   // stn[25].wipBtn[5,2] := 38000;
   // stn[25].wipBtn[5,3] := 1000;
   // stn[25].wipBtn[5,4] := 1000;
   // stn[25].wipBtn[5,5] := 1000;
   // stn[25].wipBtn[5,6] := 43000;
   // stn[25].wipBtn[5,7] := 37000;
   // stn[25].wipBtn[6,0] := 1000;
   // stn[25].wipBtn[6,1] := 244000;
   // stn[25].wipBtn[6,2] := 46000;
   // stn[25].wipBtn[6,3] := 1000;
   // stn[25].wipBtn[6,4] := 1000;
   // stn[25].wipBtn[6,5] := 1000;
   // stn[25].wipBtn[6,6] := 43000;
   // stn[25].wipBtn[6,7] := 37000;
   // stn[25].wipBtn[7,0] := 1000;
   // stn[25].wipBtn[7,1] := 244000;
   // stn[25].wipBtn[7,2] := 44000;
   // stn[25].wipBtn[7,3] := 1000;
   // stn[25].wipBtn[7,4] := 1000;
   // stn[25].wipBtn[7,5] := 1000;
   // stn[25].wipBtn[7,6] := 39000;
   // stn[25].wipBtn[7,7] := 45000;
   // stn[25].wipBtn[8,0] := 1000;
   // stn[25].wipBtn[8,1] := 244000;
   // stn[25].wipBtn[8,2] := 52000;
   // stn[25].wipBtn[8,3] := 1000;
   // stn[25].wipBtn[8,4] := 1000;
   // stn[25].wipBtn[8,5] := 1000;
   // stn[25].wipBtn[8,6] := 26000;
   // stn[25].wipBtn[8,7] := 19000;
   // stn[25].wipBtn[9,0] := 1000;
   // stn[25].wipBtn[9,1] := 244000;
   // stn[25].wipBtn[9,2] := 53000;
   // stn[25].wipBtn[9,3] := 1000;
   // stn[25].wipBtn[9,4] := 1000;
   // stn[25].wipBtn[9,5] := 1000;
   // stn[25].wipBtn[9,6] := 32000;
   // stn[25].wipBtn[9,7] := 74000;
   // stn[25].wipBtn[10,0] := 1000;
   // stn[25].wipBtn[10,1] := 244000;
   // stn[25].wipBtn[10,2] := 54000;
   // stn[25].wipBtn[10,3] := 1000;
   // stn[25].wipBtn[10,4] := 1000;
   // stn[25].wipBtn[10,5] := 1000;
   // stn[25].wipBtn[10,6] := 32000;
   // stn[25].wipBtn[10,7] := 72000;
   // stn[25].wipBtn[11,0] := 1000;
   // stn[25].wipBtn[11,1] := 244000;
   // stn[25].wipBtn[11,2] := 58000;
   // stn[25].wipBtn[11,3] := 1000;
   // stn[25].wipBtn[11,4] := 1000;
   // stn[25].wipBtn[11,5] := 1000;
   // stn[25].wipBtn[11,6] := 26000;
   // stn[25].wipBtn[11,7] := 19000;
   // stn[25].wipBtn[12,0] := 1000;
   // stn[25].wipBtn[12,1] := 244000;
   // stn[25].wipBtn[12,2] := 85000;
   // stn[25].wipBtn[12,3] := 1000;
   // stn[25].wipBtn[12,4] := 1000;
   // stn[25].wipBtn[12,5] := 1000;
   // stn[25].wipBtn[12,6] := 32000;
   // stn[25].wipBtn[12,7] := 72000;
   // stn[25].wipBtn[13,0] := 1000;
   // stn[25].wipBtn[13,1] := 244000;
   // stn[25].wipBtn[13,2] := 99000;
   // stn[25].wipBtn[13,3] := 1000;
   // stn[25].wipBtn[13,4] := 1000;
   // stn[25].wipBtn[13,5] := 1000;
   // stn[25].wipBtn[13,6] := 39000;
   // stn[25].wipBtn[13,7] := 45000;
   // stn[25].wipBtn[14,0] := 1000;
   // stn[25].wipBtn[14,1] := 244000;
   // stn[25].wipBtn[14,2] := 100000;
   // stn[25].wipBtn[14,3] := 1000;
   // stn[25].wipBtn[14,4] := 1000;
   // stn[25].wipBtn[14,5] := 1000;
   // stn[25].wipBtn[14,6] := 43000;
   // stn[25].wipBtn[14,7] := 37000;
   // stn[25].wipBtn[15,0] := 1000;
   // stn[25].wipBtn[15,1] := 244000;
   // stn[25].wipBtn[15,2] := 100000;
   // stn[25].wipBtn[15,3] := 1000;
   // stn[25].wipBtn[15,4] := 1000;
   // stn[25].wipBtn[15,5] := 1000;
   // stn[25].wipBtn[15,6] := 36000;
   // stn[25].wipBtn[15,7] := 37000;
   // stn[25].wipBtn[16,0] := 1000;
   // stn[25].wipBtn[16,1] := 244000;
   // stn[25].wipBtn[16,2] := 218000;
   // stn[25].wipBtn[16,3] := 1000;
   // stn[25].wipBtn[16,4] := 1000;
   // stn[25].wipBtn[16,5] := 1000;
   // stn[25].wipBtn[16,6] := 219000;
   // stn[25].wipBtn[16,7] := 224000;
   // stn[25].wipBtn[17,0] := 1000;
   // stn[25].wipBtn[17,1] := 244000;
   // stn[25].wipBtn[17,2] := 198000;
   // stn[25].wipBtn[17,3] := 1000;
   // stn[25].wipBtn[17,4] := 1000;
   // stn[25].wipBtn[17,5] := 1000;
   // stn[25].wipBtn[17,6] := 220000;
   // stn[25].wipBtn[17,7] := 223000;
   // stn[25].wipBtn[18,0] := 1000;
   // stn[25].wipBtn[18,1] := 244000;
   // stn[25].wipBtn[18,2] := 199000;
   // stn[25].wipBtn[18,3] := 1000;
   // stn[25].wipBtn[18,4] := 1000;
   // stn[25].wipBtn[18,5] := 1000;
   // stn[25].wipBtn[18,6] := 219000;
   // stn[25].wipBtn[18,7] := 224000;
   // stn[25].wipBtn[19,0] := 1000;
   // stn[25].wipBtn[19,1] := 244000;
   // stn[25].wipBtn[19,2] := 225000;
   // stn[25].wipBtn[19,3] := 1000;
   // stn[25].wipBtn[19,4] := 1000;
   // stn[25].wipBtn[19,5] := 1000;
   // stn[25].wipBtn[19,6] := 226000;
   // stn[25].wipBtn[19,7] := 227000;
   // stn[25].wipBtn[20,0] := 1000;
   // stn[25].wipBtn[20,1] := 244000;
   // stn[25].wipBtn[20,2] := 18000;
   // stn[25].wipBtn[20,3] := 1000;
   // stn[25].wipBtn[20,4] := 1000;
   // stn[25].wipBtn[20,5] := 1000;
   // stn[25].wipBtn[20,6] := 25000;
   // stn[25].wipBtn[20,7] := 17000;
   // stn[25].wipBtn[21,0] := 1000;
   // stn[25].wipBtn[21,1] := 244000;
   // stn[25].wipBtn[21,2] := 1000;
   // stn[25].wipBtn[21,3] := 32000;
   // stn[25].wipBtn[21,4] := 1000;
   // stn[25].wipBtn[21,5] := 1000;
   // stn[25].wipBtn[21,6] := 51000;
   // stn[25].wipBtn[21,7] := 31000;
   // stn[25].wipBtn[22,0] := 1000;
   // stn[25].wipBtn[22,1] := 244000;
   // stn[25].wipBtn[22,2] := 1000;
   // stn[25].wipBtn[22,3] := 220000;
   // stn[25].wipBtn[22,4] := 1000;
   // stn[25].wipBtn[22,5] := 1000;
   // stn[25].wipBtn[22,6] := 222000;
   // stn[25].wipBtn[22,7] := 223000;
   // stn[25].wipBtn[23,0] := 1000;
   // stn[25].wipBtn[23,1] := 244000;
   // stn[25].wipBtn[23,2] := 221000;
   // stn[25].wipBtn[23,3] := 1000;
   // stn[25].wipBtn[23,4] := 1000;
   // stn[25].wipBtn[23,5] := 1000;
   // stn[25].wipBtn[23,6] := 220000;
   // stn[25].wipBtn[23,7] := 223000;
   // stn[25].wipBtn[24,0] := 1000;
   // stn[25].wipBtn[24,1] := 1000;
   // stn[25].wipBtn[24,2] := 1000;
   // stn[25].wipBtn[24,3] := 1000;
   // stn[25].wipBtn[24,4] := 1000;
   // stn[25].wipBtn[24,5] := 1000;
   // stn[25].wipBtn[24,6] := 1000;
   // stn[25].wipBtn[24,7] := 1000;
   // stn[25].wipBtn[25,0] := 1000;
   // stn[25].wipBtn[25,1] := 1000;
   // stn[25].wipBtn[25,2] := 1000;
   // stn[25].wipBtn[25,3] := 1000;
   // stn[25].wipBtn[25,4] := 1000;
   // stn[25].wipBtn[25,5] := 1000;
   // stn[25].wipBtn[25,6] := 1000;
   // stn[25].wipBtn[25,7] := 1000;
   // stn[25].wipBtn[26,0] := 1000;
   // stn[25].wipBtn[26,1] := 1000;
   // stn[25].wipBtn[26,2] := 1000;
   // stn[25].wipBtn[26,3] := 1000;
   // stn[25].wipBtn[26,4] := 1000;
   // stn[25].wipBtn[26,5] := 1000;
   // stn[25].wipBtn[26,6] := 1000;
   // stn[25].wipBtn[26,7] := 1000;
   // stn[25].wipBtn[27,0] := 1000;
   // stn[25].wipBtn[27,1] := 1000;
   // stn[25].wipBtn[27,2] := 1000;
   // stn[25].wipBtn[27,3] := 1000;
   // stn[25].wipBtn[27,4] := 1000;
   // stn[25].wipBtn[27,5] := 1000;
   // stn[25].wipBtn[27,6] := 1000;
   // stn[25].wipBtn[27,7] := 1000;
   // stn[25].wipBtn[28,0] := 1000;
   // stn[25].wipBtn[28,1] := 1000;
   // stn[25].wipBtn[28,2] := 1000;
   // stn[25].wipBtn[28,3] := 1000;
   // stn[25].wipBtn[28,4] := 1000;
   // stn[25].wipBtn[28,5] := 1000;
   // stn[25].wipBtn[28,6] := 1000;
   // stn[25].wipBtn[28,7] := 1000;
   // stn[25].wipBtn[29,0] := 1000;
   // stn[25].wipBtn[29,1] := 1000;
   // stn[25].wipBtn[29,2] := 1000;
   // stn[25].wipBtn[29,3] := 1000;
   // stn[25].wipBtn[29,4] := 1000;
   // stn[25].wipBtn[29,5] := 1000;
   // stn[25].wipBtn[29,6] := 1000;
   // stn[25].wipBtn[29,7] := 1000;
   // stn[25].wipBtn[30,0] := 1000;
   // stn[25].wipBtn[30,1] := 1000;
   // stn[25].wipBtn[30,2] := 1000;
   // stn[25].wipBtn[30,3] := 1000;
   // stn[25].wipBtn[30,4] := 1000;
   // stn[25].wipBtn[30,5] := 1000;
   // stn[25].wipBtn[30,6] := 1000;
   // stn[25].wipBtn[30,7] := 1000;
   // stn[25].wipBtn[31,0] := 1000;
   // stn[25].wipBtn[31,1] := 1000;
   // stn[25].wipBtn[31,2] := 1000;
   // stn[25].wipBtn[31,3] := 1000;
   // stn[25].wipBtn[31,4] := 1000;
   // stn[25].wipBtn[31,5] := 1000;
   // stn[25].wipBtn[31,6] := 1000;
   // stn[25].wipBtn[31,7] := 1000;
   // stn[25].wipBtn[32,0] := 1000;
   // stn[25].wipBtn[32,1] := 1000;
   // stn[25].wipBtn[32,2] := 1000;
   // stn[25].wipBtn[32,3] := 1000;
   // stn[25].wipBtn[32,4] := 1000;
   // stn[25].wipBtn[32,5] := 1000;
   // stn[25].wipBtn[32,6] := 1000;
   // stn[25].wipBtn[32,7] := 1000;
   // stn[25].wipBtn[33,0] := 1000;
   // stn[25].wipBtn[33,1] := 1000;
   // stn[25].wipBtn[33,2] := 1000;
   // stn[25].wipBtn[33,3] := 1000;
   // stn[25].wipBtn[33,4] := 1000;
   // stn[25].wipBtn[33,5] := 1000;
   // stn[25].wipBtn[33,6] := 1000;
   // stn[25].wipBtn[33,7] := 1000;
   // stn[25].wipBtn[34,0] := 1000;
   // stn[25].wipBtn[34,1] := 1000;
   // stn[25].wipBtn[34,2] := 1000;
   // stn[25].wipBtn[34,3] := 1000;
   // stn[25].wipBtn[34,4] := 1000;
   // stn[25].wipBtn[34,5] := 1000;
   // stn[25].wipBtn[34,6] := 1000;
   // stn[25].wipBtn[34,7] := 1000;
   // stn[25].wipBtn[35,0] := 1000;
   // stn[25].wipBtn[35,1] := 1000;
   // stn[25].wipBtn[35,2] := 1000;
   // stn[25].wipBtn[35,3] := 1000;
   // stn[25].wipBtn[35,4] := 1000;
   // stn[25].wipBtn[35,5] := 1000;
   // stn[25].wipBtn[35,6] := 1000;
   // stn[25].wipBtn[35,7] := 1000;
   // stn[25].wipBtn[36,0] := 1000;
   // stn[25].wipBtn[36,1] := 1000;
   // stn[25].wipBtn[36,2] := 1000;
   // stn[25].wipBtn[36,3] := 1000;
   // stn[25].wipBtn[36,4] := 1000;
   // stn[25].wipBtn[36,5] := 1000;
   // stn[25].wipBtn[36,6] := 1000;
   // stn[25].wipBtn[36,7] := 1000;
   // stn[25].wipBtn[37,0] := 1000;
   // stn[25].wipBtn[37,1] := 1000;
   // stn[25].wipBtn[37,2] := 1000;
   // stn[25].wipBtn[37,3] := 1000;
   // stn[25].wipBtn[37,4] := 1000;
   // stn[25].wipBtn[37,5] := 1000;
   // stn[25].wipBtn[37,6] := 1000;
   // stn[25].wipBtn[37,7] := 1000;
   // stn[25].wipBtn[38,0] := 1000;
   // stn[25].wipBtn[38,1] := 1000;
   // stn[25].wipBtn[38,2] := 1000;
   // stn[25].wipBtn[38,3] := 1000;
   // stn[25].wipBtn[38,4] := 1000;
   // stn[25].wipBtn[38,5] := 1000;
   // stn[25].wipBtn[38,6] := 1000;
   // stn[25].wipBtn[38,7] := 1000;
   // stn[25].wipBtn[39,0] := 1000;
   // stn[25].wipBtn[39,1] := 1000;
   // stn[25].wipBtn[39,2] := 1000;
   // stn[25].wipBtn[39,3] := 1000;
   // stn[25].wipBtn[39,4] := 1000;
   // stn[25].wipBtn[39,5] := 1000;
   // stn[25].wipBtn[39,6] := 1000;
   // stn[25].wipBtn[39,7] := 1000;
   // stn[25].wipBtn[40,0] := 1000;
   // stn[25].wipBtn[40,1] := 1000;
   // stn[25].wipBtn[40,2] := 1000;
   // stn[25].wipBtn[40,3] := 1000;
   // stn[25].wipBtn[40,4] := 1000;
   // stn[25].wipBtn[40,5] := 1000;
   // stn[25].wipBtn[40,6] := 1000;
   // stn[25].wipBtn[40,7] := 1000;
   // stn[25].wipBtn[41,0] := 1000;
   // stn[25].wipBtn[41,1] := 1000;
   // stn[25].wipBtn[41,2] := 1000;
   // stn[25].wipBtn[41,3] := 1000;
   // stn[25].wipBtn[41,4] := 1000;
   // stn[25].wipBtn[41,5] := 1000;
   // stn[25].wipBtn[41,6] := 1000;
   // stn[25].wipBtn[41,7] := 1000;
   // stn[25].wipBtn[42,0] := 1000;
   // stn[25].wipBtn[42,1] := 1000;
   // stn[25].wipBtn[42,2] := 1000;
   // stn[25].wipBtn[42,3] := 1000;
   // stn[25].wipBtn[42,4] := 1000;
   // stn[25].wipBtn[42,5] := 1000;
   // stn[25].wipBtn[42,6] := 1000;
   // stn[25].wipBtn[42,7] := 1000;
   // stn[25].wipBtn[43,0] := 1000;
   // stn[25].wipBtn[43,1] := 1000;
   // stn[25].wipBtn[43,2] := 1000;
   // stn[25].wipBtn[43,3] := 1000;
   // stn[25].wipBtn[43,4] := 1000;
   // stn[25].wipBtn[43,5] := 1000;
   // stn[25].wipBtn[43,6] := 1000;
   // stn[25].wipBtn[43,7] := 1000;
   // stn[25].wipBtn[44,0] := 1000;
   // stn[25].wipBtn[44,1] := 1000;
   // stn[25].wipBtn[44,2] := 1000;
   // stn[25].wipBtn[44,3] := 1000;
   // stn[25].wipBtn[44,4] := 1000;
   // stn[25].wipBtn[44,5] := 1000;
   // stn[25].wipBtn[44,6] := 1000;
   // stn[25].wipBtn[44,7] := 1000;
   // stn[25].wipBtn[45,0] := 1000;
   // stn[25].wipBtn[45,1] := 1000;
   // stn[25].wipBtn[45,2] := 1000;
   // stn[25].wipBtn[45,3] := 1000;
   // stn[25].wipBtn[45,4] := 1000;
   // stn[25].wipBtn[45,5] := 1000;
   // stn[25].wipBtn[45,6] := 1000;
   // stn[25].wipBtn[45,7] := 1000;
   // stn[25].wipBtn[46,0] := 1000;
   // stn[25].wipBtn[46,1] := 1000;
   // stn[25].wipBtn[46,2] := 1000;
   // stn[25].wipBtn[46,3] := 1000;
   // stn[25].wipBtn[46,4] := 1000;
   // stn[25].wipBtn[46,5] := 1000;
   // stn[25].wipBtn[46,6] := 1000;
   // stn[25].wipBtn[46,7] := 1000;
   // stn[25].wipBtn[47,0] := 1000;
   // stn[25].wipBtn[47,1] := 1000;
   // stn[25].wipBtn[47,2] := 1000;
   // stn[25].wipBtn[47,3] := 1000;
   // stn[25].wipBtn[47,4] := 1000;
   // stn[25].wipBtn[47,5] := 1000;
   // stn[25].wipBtn[47,6] := 1000;
   // stn[25].wipBtn[47,7] := 1000;
   // stn[25].wipBtn[48,0] := 1000;
   // stn[25].wipBtn[48,1] := 1000;
   // stn[25].wipBtn[48,2] := 1000;
   // stn[25].wipBtn[48,3] := 1000;
   // stn[25].wipBtn[48,4] := 1000;
   // stn[25].wipBtn[48,5] := 1000;
   // stn[25].wipBtn[48,6] := 1000;
   // stn[25].wipBtn[48,7] := 1000;
   // stn[25].wipBtn[49,0] := 1000;
   // stn[25].wipBtn[49,1] := 1000;
   // stn[25].wipBtn[49,2] := 1000;
   // stn[25].wipBtn[49,3] := 1000;
   // stn[25].wipBtn[49,4] := 1000;
   // stn[25].wipBtn[49,5] := 1000;
   // stn[25].wipBtn[49,6] := 1000;
   // stn[25].wipBtn[49,7] := 1000;
   // stn[26].wipBtn[0,0] := 1000;
   // stn[26].wipBtn[0,1] := 244000;
   // stn[26].wipBtn[0,2] := 46000;
   // stn[26].wipBtn[0,3] := 1000;
   // stn[26].wipBtn[0,4] := 1000;
   // stn[26].wipBtn[0,5] := 1000;
   // stn[26].wipBtn[0,6] := 43000;
   // stn[26].wipBtn[0,7] := 37000;
   // stn[26].wipBtn[1,0] := 1000;
   // stn[26].wipBtn[1,1] := 244000;
   // stn[26].wipBtn[1,2] := 100000;
   // stn[26].wipBtn[1,3] := 1000;
   // stn[26].wipBtn[1,4] := 1000;
   // stn[26].wipBtn[1,5] := 1000;
   // stn[26].wipBtn[1,6] := 43000;
   // stn[26].wipBtn[1,7] := 37000;
   // stn[26].wipBtn[2,0] := 1000;
   // stn[26].wipBtn[2,1] := 244000;
   // stn[26].wipBtn[2,2] := 100000;
   // stn[26].wipBtn[2,3] := 1000;
   // stn[26].wipBtn[2,4] := 1000;
   // stn[26].wipBtn[2,5] := 1000;
   // stn[26].wipBtn[2,6] := 36000;
   // stn[26].wipBtn[2,7] := 37000;
   // stn[26].wipBtn[3,0] := 1000;
   // stn[26].wipBtn[3,1] := 244000;
   // stn[26].wipBtn[3,2] := 15000;
   // stn[26].wipBtn[3,3] := 1000;
   // stn[26].wipBtn[3,4] := 1000;
   // stn[26].wipBtn[3,5] := 16000;
   // stn[26].wipBtn[3,6] := 24000;
   // stn[26].wipBtn[3,7] := 14000;
   // stn[26].wipBtn[4,0] := 1000;
   // stn[26].wipBtn[4,1] := 244000;
   // stn[26].wipBtn[4,2] := 15000;
   // stn[26].wipBtn[4,3] := 14000;
   // stn[26].wipBtn[4,4] := 1000;
   // stn[26].wipBtn[4,5] := 48000;
   // stn[26].wipBtn[4,6] := 34000;
   // stn[26].wipBtn[4,7] := 33000;
   // stn[26].wipBtn[5,0] := 1000;
   // stn[26].wipBtn[5,1] := 244000;
   // stn[26].wipBtn[5,2] := 15000;
   // stn[26].wipBtn[5,3] := 1000;
   // stn[26].wipBtn[5,4] := 1000;
   // stn[26].wipBtn[5,5] := 16000;
   // stn[26].wipBtn[5,6] := 34000;
   // stn[26].wipBtn[5,7] := 14000;
   // stn[26].wipBtn[6,0] := 1000;
   // stn[26].wipBtn[6,1] := 244000;
   // stn[26].wipBtn[6,2] := 71000;
   // stn[26].wipBtn[6,3] := 74000;
   // stn[26].wipBtn[6,4] := 1000;
   // stn[26].wipBtn[6,5] := 59000;
   // stn[26].wipBtn[6,6] := 42000;
   // stn[26].wipBtn[6,7] := 73000;
   // stn[26].wipBtn[7,0] := 1000;
   // stn[26].wipBtn[7,1] := 244000;
   // stn[26].wipBtn[7,2] := 229000;
   // stn[26].wipBtn[7,3] := 232000;
   // stn[26].wipBtn[7,4] := 1000;
   // stn[26].wipBtn[7,5] := 230000;
   // stn[26].wipBtn[7,6] := 228000;
   // stn[26].wipBtn[7,7] := 231000;
   // stn[26].wipBtn[8,0] := 1000;
   // stn[26].wipBtn[8,1] := 244000;
   // stn[26].wipBtn[8,2] := 234000;
   // stn[26].wipBtn[8,3] := 1000;
   // stn[26].wipBtn[8,4] := 1000;
   // stn[26].wipBtn[8,5] := 230000;
   // stn[26].wipBtn[8,6] := 233000;
   // stn[26].wipBtn[8,7] := 232000;
   // stn[26].wipBtn[9,0] := 1000;
   // stn[26].wipBtn[9,1] := 244000;
   // stn[26].wipBtn[9,2] := 237000;
   // stn[26].wipBtn[9,3] := 1000;
   // stn[26].wipBtn[9,4] := 1000;
   // stn[26].wipBtn[9,5] := 238000;
   // stn[26].wipBtn[9,6] := 235000;
   // stn[26].wipBtn[9,7] := 236000;
   // stn[26].wipBtn[10,0] := 1000;
   // stn[26].wipBtn[10,1] := 244000;
   // stn[26].wipBtn[10,2] := 165000;
   // stn[26].wipBtn[10,3] := 1000;
   // stn[26].wipBtn[10,4] := 1000;
   // stn[26].wipBtn[10,5] := 166000;
   // stn[26].wipBtn[10,6] := 235000;
   // stn[26].wipBtn[10,7] := 236000;
   // stn[26].wipBtn[11,0] := 1000;
   // stn[26].wipBtn[11,1] := 244000;
   // stn[26].wipBtn[11,2] := 202000;
   // stn[26].wipBtn[11,3] := 1000;
   // stn[26].wipBtn[11,4] := 1000;
   // stn[26].wipBtn[11,5] := 201000;
   // stn[26].wipBtn[11,6] := 235000;
   // stn[26].wipBtn[11,7] := 236000;
   // stn[26].wipBtn[12,0] := 1000;
   // stn[26].wipBtn[12,1] := 244000;
   // stn[26].wipBtn[12,2] := 241000;
   // stn[26].wipBtn[12,3] := 1000;
   // stn[26].wipBtn[12,4] := 1000;
   // stn[26].wipBtn[12,5] := 242000;
   // stn[26].wipBtn[12,6] := 239000;
   // stn[26].wipBtn[12,7] := 240000;
   // stn[26].wipBtn[13,0] := 1000;
   // stn[26].wipBtn[13,1] := 244000;
   // stn[26].wipBtn[13,2] := 71000;
   // stn[26].wipBtn[13,3] := 73000;
   // stn[26].wipBtn[13,4] := 1000;
   // stn[26].wipBtn[13,5] := 59000;
   // stn[26].wipBtn[13,6] := 34000;
   // stn[26].wipBtn[13,7] := 74000;
   // stn[26].wipBtn[14,0] := 1000;
   // stn[26].wipBtn[14,1] := 1000;
   // stn[26].wipBtn[14,2] := 1000;
   // stn[26].wipBtn[14,3] := 1000;
   // stn[26].wipBtn[14,4] := 1000;
   // stn[26].wipBtn[14,5] := 1000;
   // stn[26].wipBtn[14,6] := 1000;
   // stn[26].wipBtn[14,7] := 1000;
   // stn[26].wipBtn[15,0] := 1000;
   // stn[26].wipBtn[15,1] := 1000;
   // stn[26].wipBtn[15,2] := 1000;
   // stn[26].wipBtn[15,3] := 1000;
   // stn[26].wipBtn[15,4] := 1000;
   // stn[26].wipBtn[15,5] := 1000;
   // stn[26].wipBtn[15,6] := 1000;
   // stn[26].wipBtn[15,7] := 1000;
   // stn[26].wipBtn[16,0] := 1000;
   // stn[26].wipBtn[16,1] := 1000;
   // stn[26].wipBtn[16,2] := 1000;
   // stn[26].wipBtn[16,3] := 1000;
   // stn[26].wipBtn[16,4] := 1000;
   // stn[26].wipBtn[16,5] := 1000;
   // stn[26].wipBtn[16,6] := 1000;
   // stn[26].wipBtn[16,7] := 1000;
   // stn[26].wipBtn[17,0] := 1000;
   // stn[26].wipBtn[17,1] := 1000;
   // stn[26].wipBtn[17,2] := 1000;
   // stn[26].wipBtn[17,3] := 1000;
   // stn[26].wipBtn[17,4] := 1000;
   // stn[26].wipBtn[17,5] := 1000;
   // stn[26].wipBtn[17,6] := 1000;
   // stn[26].wipBtn[17,7] := 1000;
   // stn[26].wipBtn[18,0] := 1000;
   // stn[26].wipBtn[18,1] := 1000;
   // stn[26].wipBtn[18,2] := 1000;
   // stn[26].wipBtn[18,3] := 1000;
   // stn[26].wipBtn[18,4] := 1000;
   // stn[26].wipBtn[18,5] := 1000;
   // stn[26].wipBtn[18,6] := 1000;
   // stn[26].wipBtn[18,7] := 1000;
   // stn[26].wipBtn[19,0] := 1000;
   // stn[26].wipBtn[19,1] := 1000;
   // stn[26].wipBtn[19,2] := 1000;
   // stn[26].wipBtn[19,3] := 1000;
   // stn[26].wipBtn[19,4] := 1000;
   // stn[26].wipBtn[19,5] := 1000;
   // stn[26].wipBtn[19,6] := 1000;
   // stn[26].wipBtn[19,7] := 1000;
   // stn[26].wipBtn[20,0] := 1000;
   // stn[26].wipBtn[20,1] := 1000;
   // stn[26].wipBtn[20,2] := 1000;
   // stn[26].wipBtn[20,3] := 1000;
   // stn[26].wipBtn[20,4] := 1000;
   // stn[26].wipBtn[20,5] := 1000;
   // stn[26].wipBtn[20,6] := 1000;
   // stn[26].wipBtn[20,7] := 1000;
   // stn[26].wipBtn[21,0] := 1000;
   // stn[26].wipBtn[21,1] := 1000;
   // stn[26].wipBtn[21,2] := 1000;
   // stn[26].wipBtn[21,3] := 1000;
   // stn[26].wipBtn[21,4] := 1000;
   // stn[26].wipBtn[21,5] := 1000;
   // stn[26].wipBtn[21,6] := 1000;
   // stn[26].wipBtn[21,7] := 1000;
   // stn[26].wipBtn[22,0] := 1000;
   // stn[26].wipBtn[22,1] := 1000;
   // stn[26].wipBtn[22,2] := 1000;
   // stn[26].wipBtn[22,3] := 1000;
   // stn[26].wipBtn[22,4] := 1000;
   // stn[26].wipBtn[22,5] := 1000;
   // stn[26].wipBtn[22,6] := 1000;
   // stn[26].wipBtn[22,7] := 1000;
   // stn[26].wipBtn[23,0] := 1000;
   // stn[26].wipBtn[23,1] := 1000;
   // stn[26].wipBtn[23,2] := 1000;
   // stn[26].wipBtn[23,3] := 1000;
   // stn[26].wipBtn[23,4] := 1000;
   // stn[26].wipBtn[23,5] := 1000;
   // stn[26].wipBtn[23,6] := 1000;
   // stn[26].wipBtn[23,7] := 1000;
   // stn[26].wipBtn[24,0] := 1000;
   // stn[26].wipBtn[24,1] := 1000;
   // stn[26].wipBtn[24,2] := 1000;
   // stn[26].wipBtn[24,3] := 1000;
   // stn[26].wipBtn[24,4] := 1000;
   // stn[26].wipBtn[24,5] := 1000;
   // stn[26].wipBtn[24,6] := 1000;
   // stn[26].wipBtn[24,7] := 1000;
   // stn[26].wipBtn[25,0] := 1000;
   // stn[26].wipBtn[25,1] := 1000;
   // stn[26].wipBtn[25,2] := 1000;
   // stn[26].wipBtn[25,3] := 1000;
   // stn[26].wipBtn[25,4] := 1000;
   // stn[26].wipBtn[25,5] := 1000;
   // stn[26].wipBtn[25,6] := 1000;
   // stn[26].wipBtn[25,7] := 1000;
   // stn[26].wipBtn[26,0] := 1000;
   // stn[26].wipBtn[26,1] := 1000;
   // stn[26].wipBtn[26,2] := 1000;
   // stn[26].wipBtn[26,3] := 1000;
   // stn[26].wipBtn[26,4] := 1000;
   // stn[26].wipBtn[26,5] := 1000;
   // stn[26].wipBtn[26,6] := 1000;
   // stn[26].wipBtn[26,7] := 1000;
   // stn[26].wipBtn[27,0] := 1000;
   // stn[26].wipBtn[27,1] := 1000;
   // stn[26].wipBtn[27,2] := 1000;
   // stn[26].wipBtn[27,3] := 1000;
   // stn[26].wipBtn[27,4] := 1000;
   // stn[26].wipBtn[27,5] := 1000;
   // stn[26].wipBtn[27,6] := 1000;
   // stn[26].wipBtn[27,7] := 1000;
   // stn[26].wipBtn[28,0] := 1000;
   // stn[26].wipBtn[28,1] := 1000;
   // stn[26].wipBtn[28,2] := 1000;
   // stn[26].wipBtn[28,3] := 1000;
   // stn[26].wipBtn[28,4] := 1000;
   // stn[26].wipBtn[28,5] := 1000;
   // stn[26].wipBtn[28,6] := 1000;
   // stn[26].wipBtn[28,7] := 1000;
   // stn[26].wipBtn[29,0] := 1000;
   // stn[26].wipBtn[29,1] := 1000;
   // stn[26].wipBtn[29,2] := 1000;
   // stn[26].wipBtn[29,3] := 1000;
   // stn[26].wipBtn[29,4] := 1000;
   // stn[26].wipBtn[29,5] := 1000;
   // stn[26].wipBtn[29,6] := 1000;
   // stn[26].wipBtn[29,7] := 1000;
   // stn[26].wipBtn[30,0] := 1000;
   // stn[26].wipBtn[30,1] := 1000;
   // stn[26].wipBtn[30,2] := 1000;
   // stn[26].wipBtn[30,3] := 1000;
   // stn[26].wipBtn[30,4] := 1000;
   // stn[26].wipBtn[30,5] := 1000;
   // stn[26].wipBtn[30,6] := 1000;
   // stn[26].wipBtn[30,7] := 1000;
   // stn[26].wipBtn[31,0] := 1000;
   // stn[26].wipBtn[31,1] := 1000;
   // stn[26].wipBtn[31,2] := 1000;
   // stn[26].wipBtn[31,3] := 1000;
   // stn[26].wipBtn[31,4] := 1000;
   // stn[26].wipBtn[31,5] := 1000;
   // stn[26].wipBtn[31,6] := 1000;
   // stn[26].wipBtn[31,7] := 1000;
   // stn[26].wipBtn[32,0] := 1000;
   // stn[26].wipBtn[32,1] := 1000;
   // stn[26].wipBtn[32,2] := 1000;
   // stn[26].wipBtn[32,3] := 1000;
   // stn[26].wipBtn[32,4] := 1000;
   // stn[26].wipBtn[32,5] := 1000;
   // stn[26].wipBtn[32,6] := 1000;
   // stn[26].wipBtn[32,7] := 1000;
   // stn[26].wipBtn[33,0] := 1000;
   // stn[26].wipBtn[33,1] := 1000;
   // stn[26].wipBtn[33,2] := 1000;
   // stn[26].wipBtn[33,3] := 1000;
   // stn[26].wipBtn[33,4] := 1000;
   // stn[26].wipBtn[33,5] := 1000;
   // stn[26].wipBtn[33,6] := 1000;
   // stn[26].wipBtn[33,7] := 1000;
   // stn[26].wipBtn[34,0] := 1000;
   // stn[26].wipBtn[34,1] := 1000;
   // stn[26].wipBtn[34,2] := 1000;
   // stn[26].wipBtn[34,3] := 1000;
   // stn[26].wipBtn[34,4] := 1000;
   // stn[26].wipBtn[34,5] := 1000;
   // stn[26].wipBtn[34,6] := 1000;
   // stn[26].wipBtn[34,7] := 1000;
   // stn[26].wipBtn[35,0] := 1000;
   // stn[26].wipBtn[35,1] := 1000;
   // stn[26].wipBtn[35,2] := 1000;
   // stn[26].wipBtn[35,3] := 1000;
   // stn[26].wipBtn[35,4] := 1000;
   // stn[26].wipBtn[35,5] := 1000;
   // stn[26].wipBtn[35,6] := 1000;
   // stn[26].wipBtn[35,7] := 1000;
   // stn[26].wipBtn[36,0] := 1000;
   // stn[26].wipBtn[36,1] := 1000;
   // stn[26].wipBtn[36,2] := 1000;
   // stn[26].wipBtn[36,3] := 1000;
   // stn[26].wipBtn[36,4] := 1000;
   // stn[26].wipBtn[36,5] := 1000;
   // stn[26].wipBtn[36,6] := 1000;
   // stn[26].wipBtn[36,7] := 1000;
   // stn[26].wipBtn[37,0] := 1000;
   // stn[26].wipBtn[37,1] := 1000;
   // stn[26].wipBtn[37,2] := 1000;
   // stn[26].wipBtn[37,3] := 1000;
   // stn[26].wipBtn[37,4] := 1000;
   // stn[26].wipBtn[37,5] := 1000;
   // stn[26].wipBtn[37,6] := 1000;
   // stn[26].wipBtn[37,7] := 1000;
   // stn[26].wipBtn[38,0] := 1000;
   // stn[26].wipBtn[38,1] := 1000;
   // stn[26].wipBtn[38,2] := 1000;
   // stn[26].wipBtn[38,3] := 1000;
   // stn[26].wipBtn[38,4] := 1000;
   // stn[26].wipBtn[38,5] := 1000;
   // stn[26].wipBtn[38,6] := 1000;
   // stn[26].wipBtn[38,7] := 1000;
   // stn[26].wipBtn[39,0] := 1000;
   // stn[26].wipBtn[39,1] := 1000;
   // stn[26].wipBtn[39,2] := 1000;
   // stn[26].wipBtn[39,3] := 1000;
   // stn[26].wipBtn[39,4] := 1000;
   // stn[26].wipBtn[39,5] := 1000;
   // stn[26].wipBtn[39,6] := 1000;
   // stn[26].wipBtn[39,7] := 1000;
   // stn[26].wipBtn[40,0] := 1000;
   // stn[26].wipBtn[40,1] := 1000;
   // stn[26].wipBtn[40,2] := 1000;
   // stn[26].wipBtn[40,3] := 1000;
   // stn[26].wipBtn[40,4] := 1000;
   // stn[26].wipBtn[40,5] := 1000;
   // stn[26].wipBtn[40,6] := 1000;
   // stn[26].wipBtn[40,7] := 1000;
   // stn[26].wipBtn[41,0] := 1000;
   // stn[26].wipBtn[41,1] := 1000;
   // stn[26].wipBtn[41,2] := 1000;
   // stn[26].wipBtn[41,3] := 1000;
   // stn[26].wipBtn[41,4] := 1000;
   // stn[26].wipBtn[41,5] := 1000;
   // stn[26].wipBtn[41,6] := 1000;
   // stn[26].wipBtn[41,7] := 1000;
   // stn[26].wipBtn[42,0] := 1000;
   // stn[26].wipBtn[42,1] := 1000;
   // stn[26].wipBtn[42,2] := 1000;
   // stn[26].wipBtn[42,3] := 1000;
   // stn[26].wipBtn[42,4] := 1000;
   // stn[26].wipBtn[42,5] := 1000;
   // stn[26].wipBtn[42,6] := 1000;
   // stn[26].wipBtn[42,7] := 1000;
   // stn[26].wipBtn[43,0] := 1000;
   // stn[26].wipBtn[43,1] := 1000;
   // stn[26].wipBtn[43,2] := 1000;
   // stn[26].wipBtn[43,3] := 1000;
   // stn[26].wipBtn[43,4] := 1000;
   // stn[26].wipBtn[43,5] := 1000;
   // stn[26].wipBtn[43,6] := 1000;
   // stn[26].wipBtn[43,7] := 1000;
   // stn[26].wipBtn[44,0] := 1000;
   // stn[26].wipBtn[44,1] := 1000;
   // stn[26].wipBtn[44,2] := 1000;
   // stn[26].wipBtn[44,3] := 1000;
   // stn[26].wipBtn[44,4] := 1000;
   // stn[26].wipBtn[44,5] := 1000;
   // stn[26].wipBtn[44,6] := 1000;
   // stn[26].wipBtn[44,7] := 1000;
   // stn[26].wipBtn[45,0] := 1000;
   // stn[26].wipBtn[45,1] := 1000;
   // stn[26].wipBtn[45,2] := 1000;
   // stn[26].wipBtn[45,3] := 1000;
   // stn[26].wipBtn[45,4] := 1000;
   // stn[26].wipBtn[45,5] := 1000;
   // stn[26].wipBtn[45,6] := 1000;
   // stn[26].wipBtn[45,7] := 1000;
   // stn[26].wipBtn[46,0] := 1000;
   // stn[26].wipBtn[46,1] := 1000;
   // stn[26].wipBtn[46,2] := 1000;
   // stn[26].wipBtn[46,3] := 1000;
   // stn[26].wipBtn[46,4] := 1000;
   // stn[26].wipBtn[46,5] := 1000;
   // stn[26].wipBtn[46,6] := 1000;
   // stn[26].wipBtn[46,7] := 1000;
   // stn[26].wipBtn[47,0] := 1000;
   // stn[26].wipBtn[47,1] := 1000;
   // stn[26].wipBtn[47,2] := 1000;
   // stn[26].wipBtn[47,3] := 1000;
   // stn[26].wipBtn[47,4] := 1000;
   // stn[26].wipBtn[47,5] := 1000;
   // stn[26].wipBtn[47,6] := 1000;
   // stn[26].wipBtn[47,7] := 1000;
   // stn[26].wipBtn[48,0] := 1000;
   // stn[26].wipBtn[48,1] := 1000;
   // stn[26].wipBtn[48,2] := 1000;
   // stn[26].wipBtn[48,3] := 1000;
   // stn[26].wipBtn[48,4] := 1000;
   // stn[26].wipBtn[48,5] := 1000;
   // stn[26].wipBtn[48,6] := 1000;
   // stn[26].wipBtn[48,7] := 1000;
   // stn[26].wipBtn[49,0] := 1000;
   // stn[26].wipBtn[49,1] := 1000;
   // stn[26].wipBtn[49,2] := 1000;
   // stn[26].wipBtn[49,3] := 1000;
   // stn[26].wipBtn[49,4] := 1000;
   // stn[26].wipBtn[49,5] := 1000;
   // stn[26].wipBtn[49,6] := 1000;
   // stn[26].wipBtn[49,7] := 1000;
   // stn[27].wipBtn[0,0] := 1000;
   // stn[27].wipBtn[0,1] := 244000;
   // stn[27].wipBtn[0,2] := 149000;
   // stn[27].wipBtn[0,3] := 1000;
   // stn[27].wipBtn[0,4] := 1000;
   // stn[27].wipBtn[0,5] := 1000;
   // stn[27].wipBtn[0,6] := 148000;
   // stn[27].wipBtn[0,7] := 150000;
   // stn[27].wipBtn[1,0] := 1000;
   // stn[27].wipBtn[1,1] := 244000;
   // stn[27].wipBtn[1,2] := 54000;
   // stn[27].wipBtn[1,3] := 1000;
   // stn[27].wipBtn[1,4] := 1000;
   // stn[27].wipBtn[1,5] := 1000;
   // stn[27].wipBtn[1,6] := 32000;
   // stn[27].wipBtn[1,7] := 72000;
   // stn[27].wipBtn[2,0] := 1000;
   // stn[27].wipBtn[2,1] := 244000;
   // stn[27].wipBtn[2,2] := 58000;
   // stn[27].wipBtn[2,3] := 1000;
   // stn[27].wipBtn[2,4] := 1000;
   // stn[27].wipBtn[2,5] := 1000;
   // stn[27].wipBtn[2,6] := 26000;
   // stn[27].wipBtn[2,7] := 19000;
   // stn[27].wipBtn[3,0] := 1000;
   // stn[27].wipBtn[3,1] := 244000;
   // stn[27].wipBtn[3,2] := 85000;
   // stn[27].wipBtn[3,3] := 1000;
   // stn[27].wipBtn[3,4] := 1000;
   // stn[27].wipBtn[3,5] := 1000;
   // stn[27].wipBtn[3,6] := 32000;
   // stn[27].wipBtn[3,7] := 72000;
   // stn[27].wipBtn[4,0] := 1000;
   // stn[27].wipBtn[4,1] := 244000;
   // stn[27].wipBtn[4,2] := 71000;
   // stn[27].wipBtn[4,3] := 73000;
   // stn[27].wipBtn[4,4] := 1000;
   // stn[27].wipBtn[4,5] := 59000;
   // stn[27].wipBtn[4,6] := 34000;
   // stn[27].wipBtn[4,7] := 74000;
   // stn[27].wipBtn[5,0] := 1000;
   // stn[27].wipBtn[5,1] := 244000;
   // stn[27].wipBtn[5,2] := 128000;
   // stn[27].wipBtn[5,3] := 1000;
   // stn[27].wipBtn[5,4] := 1000;
   // stn[27].wipBtn[5,5] := 101000;
   // stn[27].wipBtn[5,6] := 102000;
   // stn[27].wipBtn[5,7] := 129000;
   // stn[27].wipBtn[6,0] := 1000;
   // stn[27].wipBtn[6,1] := 244000;
   // stn[27].wipBtn[6,2] := 123000;
   // stn[27].wipBtn[6,3] := 124000;
   // stn[27].wipBtn[6,4] := 1000;
   // stn[27].wipBtn[6,5] := 103000;
   // stn[27].wipBtn[6,6] := 104000;
   // stn[27].wipBtn[6,7] := 134000;
   // stn[27].wipBtn[7,0] := 1000;
   // stn[27].wipBtn[7,1] := 244000;
   // stn[27].wipBtn[7,2] := 101000;
   // stn[27].wipBtn[7,3] := 129000;
   // stn[27].wipBtn[7,4] := 1000;
   // stn[27].wipBtn[7,5] := 103000;
   // stn[27].wipBtn[7,6] := 105000;
   // stn[27].wipBtn[7,7] := 134000;
   // stn[27].wipBtn[8,0] := 1000;
   // stn[27].wipBtn[8,1] := 244000;
   // stn[27].wipBtn[8,2] := 106000;
   // stn[27].wipBtn[8,3] := 124000;
   // stn[27].wipBtn[8,4] := 1000;
   // stn[27].wipBtn[8,5] := 107000;
   // stn[27].wipBtn[8,6] := 108000;
   // stn[27].wipBtn[8,7] := 134000;
   // stn[27].wipBtn[9,0] := 1000;
   // stn[27].wipBtn[9,1] := 244000;
   // stn[27].wipBtn[9,2] := 101000;
   // stn[27].wipBtn[9,3] := 1000;
   // stn[27].wipBtn[9,4] := 1000;
   // stn[27].wipBtn[9,5] := 128000;
   // stn[27].wipBtn[9,6] := 108000;
   // stn[27].wipBtn[9,7] := 129000;
   // stn[27].wipBtn[10,0] := 1000;
   // stn[27].wipBtn[10,1] := 244000;
   // stn[27].wipBtn[10,2] := 101000;
   // stn[27].wipBtn[10,3] := 129000;
   // stn[27].wipBtn[10,4] := 1000;
   // stn[27].wipBtn[10,5] := 107000;
   // stn[27].wipBtn[10,6] := 108000;
   // stn[27].wipBtn[10,7] := 124000;
   // stn[27].wipBtn[11,0] := 1000;
   // stn[27].wipBtn[11,1] := 244000;
   // stn[27].wipBtn[11,2] := 109000;
   // stn[27].wipBtn[11,3] := 1000;
   // stn[27].wipBtn[11,4] := 1000;
   // stn[27].wipBtn[11,5] := 1000;
   // stn[27].wipBtn[11,6] := 108000;
   // stn[27].wipBtn[11,7] := 110000;
   // stn[27].wipBtn[12,0] := 1000;
   // stn[27].wipBtn[12,1] := 244000;
   // stn[27].wipBtn[12,2] := 111000;
   // stn[27].wipBtn[12,3] := 114000;
   // stn[27].wipBtn[12,4] := 1000;
   // stn[27].wipBtn[12,5] := 113000;
   // stn[27].wipBtn[12,6] := 115000;
   // stn[27].wipBtn[12,7] := 112000;
   // stn[27].wipBtn[13,0] := 1000;
   // stn[27].wipBtn[13,1] := 244000;
   // stn[27].wipBtn[13,2] := 116000;
   // stn[27].wipBtn[13,3] := 1000;
   // stn[27].wipBtn[13,4] := 1000;
   // stn[27].wipBtn[13,5] := 113000;
   // stn[27].wipBtn[13,6] := 115000;
   // stn[27].wipBtn[13,7] := 114000;
   // stn[27].wipBtn[14,0] := 1000;
   // stn[27].wipBtn[14,1] := 244000;
   // stn[27].wipBtn[14,2] := 117000;
   // stn[27].wipBtn[14,3] := 112000;
   // stn[27].wipBtn[14,4] := 1000;
   // stn[27].wipBtn[14,5] := 119000;
   // stn[27].wipBtn[14,6] := 115000;
   // stn[27].wipBtn[14,7] := 118000;
   // stn[27].wipBtn[15,0] := 1000;
   // stn[27].wipBtn[15,1] := 244000;
   // stn[27].wipBtn[15,2] := 117000;
   // stn[27].wipBtn[15,3] := 118000;
   // stn[27].wipBtn[15,4] := 1000;
   // stn[27].wipBtn[15,5] := 119000;
   // stn[27].wipBtn[15,6] := 121000;
   // stn[27].wipBtn[15,7] := 112000;
   // stn[27].wipBtn[16,0] := 1000;
   // stn[27].wipBtn[16,1] := 244000;
   // stn[27].wipBtn[16,2] := 120000;
   // stn[27].wipBtn[16,3] := 1000;
   // stn[27].wipBtn[16,4] := 1000;
   // stn[27].wipBtn[16,5] := 122000;
   // stn[27].wipBtn[16,6] := 115000;
   // stn[27].wipBtn[16,7] := 112000;
   // stn[27].wipBtn[17,0] := 1000;
   // stn[27].wipBtn[17,1] := 244000;
   // stn[27].wipBtn[17,2] := 125000;
   // stn[27].wipBtn[17,3] := 126000;
   // stn[27].wipBtn[17,4] := 1000;
   // stn[27].wipBtn[17,5] := 123000;
   // stn[27].wipBtn[17,6] := 108000;
   // stn[27].wipBtn[17,7] := 124000;
   // stn[27].wipBtn[18,0] := 1000;
   // stn[27].wipBtn[18,1] := 244000;
   // stn[27].wipBtn[18,2] := 101000;
   // stn[27].wipBtn[18,3] := 1000;
   // stn[27].wipBtn[18,4] := 1000;
   // stn[27].wipBtn[18,5] := 128000;
   // stn[27].wipBtn[18,6] := 127000;
   // stn[27].wipBtn[18,7] := 129000;
   // stn[27].wipBtn[19,0] := 1000;
   // stn[27].wipBtn[19,1] := 244000;
   // stn[27].wipBtn[19,2] := 128000;
   // stn[27].wipBtn[19,3] := 124000;
   // stn[27].wipBtn[19,4] := 1000;
   // stn[27].wipBtn[19,5] := 123000;
   // stn[27].wipBtn[19,6] := 130000;
   // stn[27].wipBtn[19,7] := 129000;